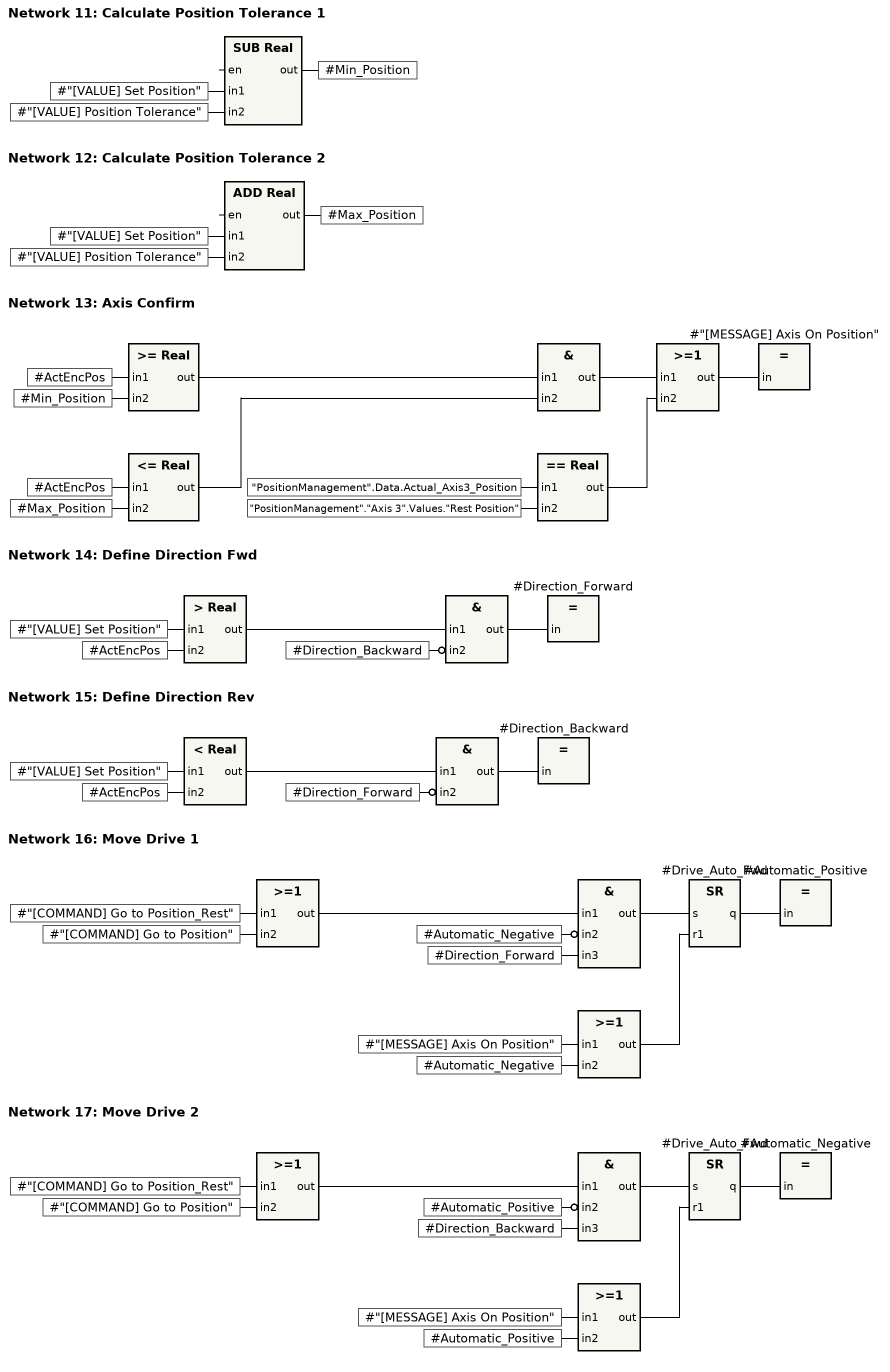
   #Min_Position := #"[VALUE] Set Position" - #"[VALUE] Position Tolerance";
END_REGION

REGION Network 12: Calculate Position Tolerance 2
   #Max_Position := #"[VALUE] Set Position" + #"[VALUE] Position Tolerance";
END_REGION

REGION Network 13: Axis Confirm
   #"[MESSAGE] Axis On Position" := ((#ActEncPos >= #Min_Position) AND (#ActEncPos <= #Max_Position)) OR ("PositionManagement".Data.Actual_Axis3_Position = "PositionManagement"."Axis 3".Values."Rest Position");
END_REGION

REGION Network 14: Define Direction Fwd
   #Direction_Forward := (#"[VALUE] Set Position" > #ActEncPos) AND NOT #Direction_Backward;
END_REGION

REGION Network 15: Define Direction Rev
   #Direction_Backward := (#"[VALUE] Set Position" < #ActEncPos) AND NOT #Direction_Forward;
END_REGION

REGION Network 16: Move Drive 1
   IF (#"[COMMAND] Go to Position_Rest" OR #"[COMMAND] Go to Position") AND NOT #Automatic_Negative AND #Direction_Forward THEN
       #Drive_Auto_Fwd := TRUE;   // SR flip-flop
   END_IF;
   IF #"[MESSAGE] Axis On Position" OR #Automatic_Negative THEN #Drive_Auto_Fwd := FALSE; END_IF;
   #Automatic_Positive := #Drive_Auto_Fwd;
END_REGION

REGION Network 17: Move Drive 2
   IF (#"[COMMAND] Go to Position_Rest" OR #"[COMMAND] Go to Position") AND NOT #Automatic_Positive AND #Direction_Backward THEN
       #Drive_Auto_Fwd := TRUE;   // SR flip-flop
   END_IF;
   IF #"[MESSAGE] Axis On Position" OR #Automatic_Positive THEN #Drive_Auto_Fwd := FALSE; END_IF;
   #Automatic_Negative := #Drive_Auto_Fwd;
END_REGION

REGION Network 18: Manual Displacement Positive
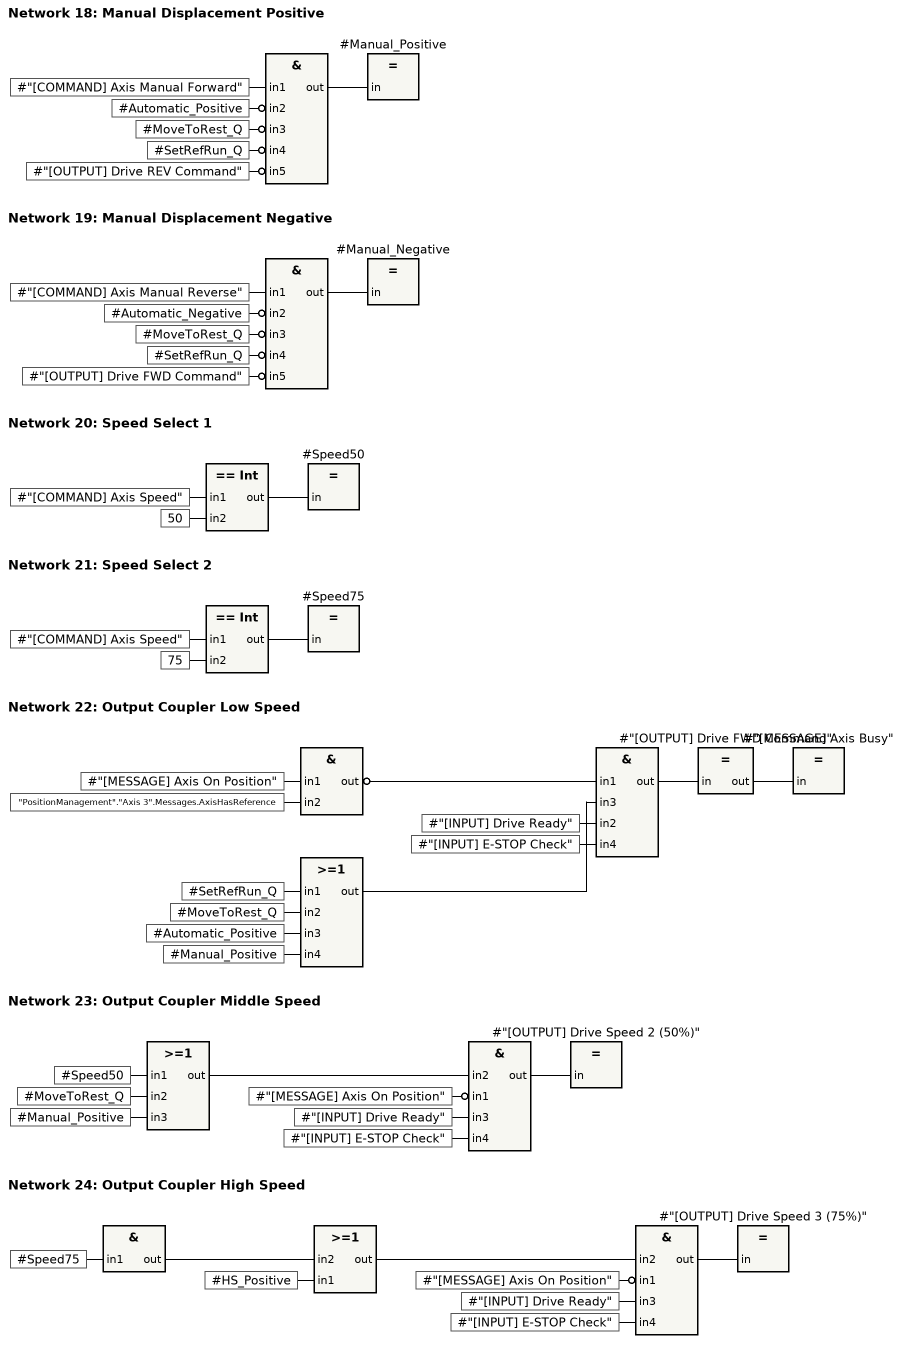
   #Manual_Positive := #"[COMMAND] Axis Manual Forward" AND NOT #Automatic_Positive AND NOT #MoveToRest_Q AND NOT #SetRefRun_Q AND NOT #"[OUTPUT] Drive REV Command";
END_REGION

REGION Network 19: Manual Displacement Negative
   #Manual_Negative := #"[COMMAND] Axis Manual Reverse" AND NOT #Automatic_Negative AND NOT #MoveToRest_Q AND NOT #SetRefRun_Q AND NOT #"[OUTPUT] Drive FWD Command";
END_REGION

REGION Network 20: Speed Select 1
   #Speed50 := #"[COMMAND] Axis Speed" = 50;
END_REGION

REGION Network 21: Speed Select 2
   #Speed75 := #"[COMMAND] Axis Speed" = 75;
END_REGION

REGION Network 22: Output Coupler Low Speed
   #_w1 := NOT (#"[MESSAGE] Axis On Position" AND "PositionManagement"."Axis 3".Messages.AxisHasReference) AND (#SetRefRun_Q OR #MoveToRest_Q OR #Automatic_Positive OR #Manual_Positive) AND #"[INPUT] Drive Ready" AND #"[INPUT] E-STOP Check";
   #"[OUTPUT] Drive FWD Command" := #_w1;
   #"[MESSAGE] Axis Busy" := #_w1;
END_REGION

REGION Network 23: Output Coupler Middle Speed
   #"[OUTPUT] Drive Speed 2 (50%)" := (#Speed50 OR #MoveToRest_Q OR #Manual_Positive) AND NOT #"[MESSAGE] Axis On Position" AND #"[INPUT] Drive Ready" AND #"[INPUT] E-STOP Check";
END_REGION

REGION Network 24: Output Coupler High Speed
   #"[OUTPUT] Drive Speed 3 (75%)" := (#Speed75 OR #HS_Positive) AND NOT #"[MESSAGE] Axis On Position" AND #"[INPUT] Drive Ready" AND #"[INPUT] E-STOP Check";
END_REGION

REGION Network 25: Output Coupler Reverse
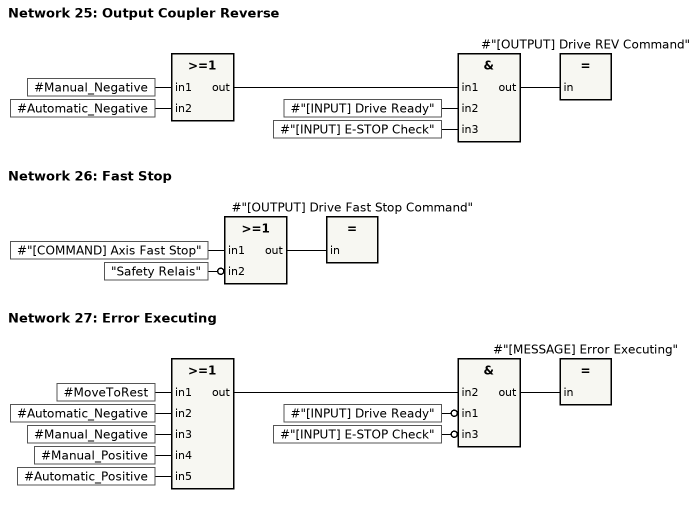
   #"[OUTPUT] Drive REV Command" := (#Manual_Negative OR #Automatic_Negative) AND #"[INPUT] Drive Ready" AND #"[INPUT] E-STOP Check";
END_REGION

REGION Network 26: Fast Stop
   #"[OUTPUT] Drive Fast Stop Command" := #"[COMMAND] Axis Fast Stop" OR NOT "Safety Relais";
END_REGION

REGION Network 27: Error Executing
   #"[MESSAGE] Error Executing" := (#MoveToRest OR #Automatic_Negative OR #Manual_Negative OR #Manual_Positive OR #Automatic_Positive) AND NOT #"[INPUT] Drive Ready" AND NOT #"[INPUT] E-STOP Check";
END_REGION
END_FUNCTION

(* ===== HMI "HMI_RT_2" =====
system functions are stored by id; their names below are inferred from use
connection "HMI_Connection_1": ETHERNET, SIMATIC S7 300/400 MPI

HMI tags "Default tag table"
   "Tag_ScreenNumber" : UInt, internal
   "Alle uitgangen(1)" : Bool = PLC "Alle uitgangen(1)" AT %I1.4, 1 s
   "Product op de band" : Bool = PLC "Sensor Op Band" AT %I0.6, 1 s
   "Product op de band(1)" : Bool = PLC "Sensor Op Band" AT %I0.6, 1 s
   "Trechter moet worden bijgevuld" : Bool = PLC "Sensor Trechter" AT %I0.5, 1 s
   "Voorverdeelwals staat in positie" : Bool = PLC "Sensor Wals (Option)" AT %I0.7, 1 s
   "Programma 1 draaid" : Bool = PLC "Programma 1" AT %I2.0, 1 s
   "Programma 2 draaid" : Bool = PLC "Programma 2" AT %I2.1, 1 s
   "Progrmma 3 draaid" : Bool = PLC "Programma 3" AT %I2.2, 1 s
   "Machine staat aan" : Bool = PLC "Start Machine" AT %I2.4, 1 s
   "Machine staat ui" : Bool = PLC "Stop Machine" AT %I2.5, 1 s
   "Noodstop machine" : Bool = PLC "ESB Pressend" AT %I1.1, 1 s
   "Startknop_Scherm" : Bool = PLC Startknop_Scherm AT %M15.0, 1 s
   "Stopknop_Scherm" : Bool = PLC Stopknop_Scherm AT %M15.1, 1 s
   "Systeem RUN" : Bool = PLC "Systeem RUN" AT %M0.0, 1 s
   "Reset Active" : Bool = PLC "Reset Active" AT %I1.2, 1 s
   "Drive 1 Ready" : Bool = PLC "Drive 1 Ready" AT %I0.0, 1 s
   "Drive 2 Ready" : Bool = PLC "Drive 2 Ready" AT %I0.1, 1 s
   "Drive 3 Ready" : Bool = PLC "Drive 3 Ready" AT %I0.2, 1 s
   "Drive 4 Ready" : Bool = PLC "Drive 4 Ready" AT %I0.3, 1 s
   "Drive 5 Ready" : Bool = PLC "Drive 5 Ready" AT %I0.4, 1 s
   "Drive 2 RUN FWD" : Bool = PLC "Drive 2 RUN FWD" AT %Q1.5, 1 s
   "Drive 1 RUN FWD" : Bool = PLC "Drive 1 RUN FWD" AT %Q1.0, 1 s
   "Drive 1 Speed 1" : Bool = PLC "Drive 1 Speed 1" AT %Q1.2, 1 s
   "Drive 1 Speed 2" : Bool = PLC "Drive 1 Speed 2" AT %Q1.3, 1 s
   "Drive 3 RUN FWD" : Bool = PLC "Drive 3 RUN FWD" AT %Q2.2, 1 s
   "Valve 1" : Bool = PLC "Valve 1" AT %Q4.6, 1 s
   "Drive 4 RUN FWD" : Bool = PLC "Drive 4 RUN FWD" AT %Q2.7, 1 s
   "StopAll" : Bool = PLC StopAll AT %M20.4, 1 s
   "Safety Relais" : Bool = PLC "Safety Relais" AT %Q0.0, 1 s
   "Drive_1_Manual" : Bool = PLC Drive_1_Manual AT %M50.1, 1 s
   "Stop_drive_1" : Bool = PLC Stop_drive_1 AT %M52.4, 1 s
   "Drive_2_Manual" : Bool = PLC Drive_2_Manual AT %M50.3, 1 s
   "Stop_drive_2" : Bool = PLC Stop_drive_2 AT %M52.5, 1 s
   "Drive_3_Manual" : Bool = PLC Drive_3_Manual AT %M50.5, 1 s
   "Stop_drive_3" : Bool = PLC Stop_drive_3 AT %M52.6, 1 s
   "Valve_1_Manual" : Bool = PLC Valve_1_Manual AT %M51.3, 1 s
   "Drive_4_Manual" : Bool = PLC Drive_4_Manual AT %M50.7, 1 s
   "Drive_5_Manual" : Bool = PLC Drive_5_Manual AT %M51.1, 1 s
   "Trechter_Bijvullen_Signaal" : Bool = PLC Trechter_Bijvullen_Signaal AT %M53.6, 1 s
   "RUN_Manual" : Bool = PLC RUN_Manual AT %M101.0, 1 s
   "Safety_Override" : Bool = PLC Safety_Override AT %M100.6, 1 s
   "Invert_Trechter_Sensor" : Bool = PLC Invert_Trechter_Sensor AT %M101.2, 1 s
   "Drive 1 REV]" : Bool = PLC "Drive 1 REV]" AT %Q1.1, 1 s
   "Drive 1 Rapid Stop" : Bool = PLC "Drive 1 Rapid Stop" AT %Q0.3, 1 s
   "Drive 2 Rapid Stop" : Bool = PLC "Drive 2 Rapid Stop" AT %Q0.4, 1 s
   "Drive 2 REV" : Bool = PLC "Drive 2 REV" AT %Q1.6, 1 s
   "Drive 3 Rapid Stop" : Bool = PLC "Drive 3 Rapid Stop" AT %Q0.5, 1 s
   "Drive 3 REV" : Bool = PLC "Drive 3 REV" AT %Q2.3, 1 s
   "Disable_Module" : Bool = PLC Disable_Module AT %M101.4, 1 s
   "PLCMemory_Safety_Delay" : Time = PLC PLCMemory.Safety_Delay AT %DB15.DBD8, 1 s
   "PLCMemory_Magazijn_Sensor_Delay" : Time = PLC PLCMemory.Offset_Timers.Magazijn_Sensor_Delay AT %DB15.DBD600, 1 s
   "PLCMemory_Homing_Sensor_Wals_Offset_Test" : Time = PLC PLCMemory.Homing_Sensor_Wals_Offset_Test AT %DB15.DBD0, 1 s
   "PLCMemory_Wals_Delay_Offset" : Time = PLC PLCMemory.Wals_Delay_Offset AT %DB15.DBD4, 1 s
   "PLCMemory_Aanvoer_Start_Offset" : Time = PLC PLCMemory.Offset_Timers.Aanvoer_Start_Offset AT %DB15.DBD596, 1 s
   "PLCMemory_Aanvoer_Stop_Offset" : Time = PLC PLCMemory.Offset_Timers.Aanvoer_Stop_Offset AT %DB15.DBD604, 1 s
   "PLCMemory_Trilgoten_Start_Offset" : Time = PLC PLCMemory.Offset_Timers.Trilgoten_Start_Offset AT %DB15.DBD588, 1 s
   "PLCMemory_Trilgoten_Stop_Offset" : Time = PLC PLCMemory.Offset_Timers.Trilgoten_Stop_Offset AT %DB15.DBD592, 1 s
   "Alarm_Axis_Not_Position" : Bool = PLC Alarm_Axis_Not_Position AT %M54.1, 1 s
   "PLCMemory_WalsCheck_Time" : Time = PLC PLCMemory.WalsCheck_Time AT %DB15.DBD12, 1 s
   "Alarm_Product_Not_Position" : Bool = PLC Alarm_Product_Not_Position AT %M54.2, 1 s
   "PLCMemory_ProductCheck_Time" : Time = PLC PLCMemory.ProductCheck_Time AT %DB15.DBD16, 1 s
   "LED Programma 1" : Bool = PLC "LED Programma 1" AT %Q4.1, 1 s
   "LED Programma 2" : Bool = PLC "LED Programma 2" AT %Q4.2, 1 s
   "LED Programma 3" : Bool = PLC "LED Programma 3" AT %Q4.3, 1 s
   "PLCMemory_ProductIntervalTime" : Time = PLC PLCMemory.ProductIntervalTime AT %DB15.DBD20, 1 s
   "PLCMemory_TD_Products_Counter" : Int = PLC PLCMemory.TD_Products_Counter AT %DB15.DBW32, 1 s
   "ResetTotalProducts" : Bool = PLC ResetTotalProducts AT %M102.7, 1 s
   "Door_Safety_Alarm" : Bool = PLC Door_Safety_Alarm AT %M54.3, 1 s
   "ESB_Safety_Alarm" : Bool = PLC ESB_Safety_Alarm AT %M54.4, 1 s
   "Valve_2_Manual" : Bool = PLC Valve_2_Manual AT %M51.5, 1 s
   "Valve 2" : Bool = PLC "Valve 2" AT %Q4.7, 1 s
   "Cilinder Trechterwissel in" : Bool = PLC "Spare(5)" AT %I3.0, 1 s
   "Cilinder Trechterwissel uit" : Bool = PLC "Spare(6)" AT %I3.1, 1 s
   "Valve 3" : Bool = PLC "Valve 3" AT %Q5.0, 1 s
   "Valve 4" : Bool = PLC "Valve 4" AT %Q5.1, 1 s
   "Valve 5" : Bool = PLC "Valve 5" AT %Q5.2, 1 s
   "Valve_3_Manual" : Bool = PLC Valve_3_Manual AT %M51.7, 1 s
   "Valve_4_Manual" : Bool = PLC Valve_4_Manual AT %M52.1, 1 s
   "Valve_5_Manual" : Bool = PLC Valve_5_Manual AT %M52.3, 1 s
   "Drive 5 REV" : Bool = PLC "Drive 5 REV" AT %Q3.5, 1 s
   "Drive 5 RUN FWD" : Bool = PLC "Drive 5 RUN FWD" AT %Q3.4, 1 s
   "Drive 5 Rapid Stop" : Bool = PLC "Drive 5 Rapid Stop" AT %Q0.7, 1 s
   "ESB Oke" : Bool = PLC "ESB Oke" AT %I1.0, 1 s
   "Door 1 NC contact" : Bool = PLC "Door 1 NC contact" AT %I1.5, 1 s
   "Door 2 NC contact" : Bool = PLC "Door 2 NC contact" AT %I1.7, 1 s
   "Sensor_op_band_memory" : Bool = PLC Sensor_op_band_memory AT %M15.3, 1 s
   "Drive_3_Auto" : Bool = PLC Drive_3_Auto AT %M50.4, 1 s
   "WalsSensorMemory" : Bool = PLC WalsSensorMemory AT %M101.3, 1 s
   "Drive_2_Auto" : Bool = PLC Drive_2_Auto AT %M50.2, 1 s
   "Drive_1_Auto" : Bool = PLC Drive_1_Auto AT %M50.0, 1 s
   "Alarms_AlarmsWord" : Word = PLC Alarms.AlarmsWord AT %DB24.DBW2, 1 s
   "Clear_Error" : Int, internal
   "Alarms_AlarmStruct_Alarm_Drive1" : Bool = PLC Alarms.AlarmStruct.Alarm_Drive1 AT %DB24.DBX0.2, 1 s
   "Alarms_HMI_Alarm_Drive1" : Word = PLC Alarms.HMI_Alarm_Drive1 AT %DB24.DBW4, 1 s
   "Alarms_HMI_Alarm_Drive2" : Word = PLC Alarms.HMI_Alarm_Drive2 AT %DB24.DBW6, 1 s
   "Alarms_HMI_Alarm_Drive3" : Word = PLC Alarms.HMI_Alarm_Drive3 AT %DB24.DBW8, 1 s
   "Alarms_HMI_Alarm_Drive4" : Word = PLC Alarms.HMI_Alarm_Drive4 AT %DB24.DBW10, 1 s
   "Alarms_HMI_Alarm_Drive5" : Word = PLC Alarms.HMI_Alarm_Drive5 AT %DB24.DBW12, 1 s
   "Sleutelschakelaar_Ingang" : Bool = PLC "Noodsleutel(1)" AT %I1.3, 1 s
      on ChangeValue: function_a9b89908("PLCMemory_UsernameMemory", "PLCMemory_PasswordMemory")
   "PLCMemory_UsernameMemory" : String[254] = PLC PLCMemory.UsernameMemory AT %DB15.DBX34.0, 1 s
   "PLCMemory_PasswordMemory" : String[254] = PLC PLCMemory.PasswordMemory AT %DB15.DBX290.0, 1 s
   "Drive 4 REV" : Bool = PLC "Drive 4 REV" AT %Q3.0, 1 s
   "Drive 4 Rapid Stop" : Bool = PLC "Drive 4 Rapid Stop" AT %Q0.6, 1 s
   "PLCMemory_SpeedSettingsTakeover" : Bool = PLC PLCMemory.SpeedSettingsTakeover AT %DB15.DBX546.0, 1 s
   "PLCMemory_SpeedSettingBand" : Bool = PLC PLCMemory.SpeedSettingBand AT %DB15.DBX546.2, 1 s
   "PLCMemory_TimingSettingOvername" : Bool = PLC PLCMemory.TimingSettingOvername AT %DB15.DBX546.3, 1 s
   "PLCMemory_SpeedSettingOvername" : Bool = PLC PLCMemory.SpeedSettingOvername AT %DB15.DBX546.1, 1 s
   "PLCMemory_Overname_Start_Offset" : Time = PLC PLCMemory.Offset_Timers.Overname_Start_Offset AT %DB15.DBD608, 1 s
   "PLCMemory_Overname_Stop_Offset" : Time = PLC PLCMemory.Offset_Timers.Overname_Stop_Offset AT %DB15.DBD612, 1 s
   "PLCMemory_EncoderPosition" : Real = PLC PLCMemory.EncoderPosition AT %DB15.DBD548, 1 s
   "PLCMemory_StepSize" : Real = PLC PLCMemory.StepSize AT %DB15.DBD552, 1 s
   "PLCMemory_Desired_Encoder_Position" : Real = PLC PLCMemory.Desired_Encoder_Position AT %DB15.DBD556, 1 s
   "HMI_Des_Pos_Axis3" : Bool = PLC HMI_Des_Pos_Axis3 AT %M54.5, 1 s
   "PLCMemory_Encoder PulsOffset" : Time = PLC PLCMemory."Encoder PulsOffset" AT %DB15.DBD564, 1 s
   "PLCMemory_Tolerance" : Real = PLC PLCMemory.Tolerance AT %DB15.DBD560, 1 s
   "PLCMemory_Axis3_Ref_Pos" : Real = PLC PLCMemory.Axis3_Ref_Pos AT %DB15.DBD568, 1 s
   "Cleaning_Active" : Bool = PLC Cleaning_Active AT %M182.0, 1 s
   "Cleaning" : Bool = PLC Cleaning AT %I2.3, 1 s
   "Cleaning_Confirmed" : Bool = PLC Cleaning_Confirmed AT %M182.1, 1 s
   "Cleaning_Cancelled" : Bool = PLC Cleaning_Cancelled AT %M182.2, 1 s
   "Cleaning_Screen_Active" : Bool = PLC Cleaning_Screen_Active AT %M182.3, 1 s
   "Tag_19" : Bool = PLC Tag_19 AT %M160.0, 1 s
   "Safety_Doors" : Bool = PLC Safety_Doors AT %M112.2, 1 s
   "HMI_ManualControl" : Bool = PLC HMI_ManualControl AT %M182.5, 1 s
   "PositionManagement_Data_Actual_Axis1_Position" : Real = PLC PositionManagement.Data.Actual_Axis3_Position AT %DB51.DBD16, 100 ms
   "PositionManagement_Axis 3_Values_Set Position" : Real, internal
   "PositionManagement_Axis 3_Commands_Go To Position" : Bool = PLC PositionManagement."Axis 3".Commands."Go To Position" AT %DB51.DBX312.3, 1 s
   "PositionManagement_Axis 3_Values_Pulsfactor" : Real = PLC PositionManagement."Axis 3".Values.Pulsfactor AT %DB51.DBD306, 1 s
   "PositionManagement_Axis 3_Values_Position Offset" : Real = PLC PositionManagement."Axis 3".Values."Position Offset" AT %DB51.DBD302, 1 s
   "PositionManagement_Axis 3_Values_Reference Position" : Int = PLC PositionManagement."Axis 3".Values."Reference Position" AT %DB51.DBW280, 1 s
   "PositionManagement_Axis 3_Values_Rest Position" : Real = PLC PositionManagement."Axis 3".Values."Rest Position" AT %DB51.DBD286, 1 s
   "PositionManagement_Axis 3_Values_Axis Correction" : Real = PLC PositionManagement."Axis 3".Values."Axis Correction" AT %DB51.DBD298, 1 s
   "PositionManagement_Axis 3_Values_Axis_Speed" : Int = PLC PositionManagement."Axis 3".Values.Axis_Speed AT %DB51.DBW310, 1 s
   "Drive_3_Manual_Rev" : Bool = PLC Drive_3_Manual_Rev AT %M60.1, 1 s
   "Manual Jog Fwd" : Bool = PLC "Manual Jog Fwd" AT %M137.0, 1 s
   "Manual Jog Rev" : Bool = PLC "Manual Jog Rev" AT %M137.1, 1 s
   "Counter2_IW102" : Int = PLC Counter2_IW102 AT %IW102, 1 s
   "PositionManagement_Axis 3_Commands_Start Ref Run" : Bool = PLC PositionManagement."Axis 3".Commands."Start Ref Run" AT %DB51.DBX312.1, 1 s
   "PLCMemory_Disable_Modules_Disable_Aandruk1" : Bool = PLC PLCMemory.Disable_Modules.Disable_Aandruk1 AT %DB15.DBX586.3, 1 s
   "PLCMemory_Disable_Modules_Disable_Aandruk2" : Bool = PLC PLCMemory.Disable_Modules.Disable_Aandruk2 AT %DB15.DBX586.4, 1 s
   "PLCMemory_Disable_Modules_Disable_Aandruk3" : Bool = PLC PLCMemory.Disable_Modules.Disable_Aandruk3 AT %DB15.DBX586.5, 1 s
   "PLCMemory_Disable_Modules_Disable_Blaaspuls" : Bool = PLC PLCMemory.Disable_Modules.Disable_Blaaspuls AT %DB15.DBX586.6, 1 s
   "PLCMemory_Disable_Modules_Disable_Afsluiter" : Bool = PLC PLCMemory.Disable_Modules.Disable_Afsluiter AT %DB15.DBX587.0, 1 s
   "PLCMemory_Offset_Timers_BlowOff_CycleTime" : Time = PLC PLCMemory.Offset_Timers.BlowOff_CycleTime AT %DB15.DBD624, 1 s
   "PLCMemory_Offset_Timers_Blow_Off_PulseTime" : Time = PLC PLCMemory.Offset_Timers.Blow_Off_PulseTime AT %DB15.DBD628, 1 s
   "PLCMemory_Disable_Modules_Disable_Retourband" : Bool = PLC PLCMemory.Disable_Modules.Disable_Retourband AT %DB15.DBX586.7, 1 s
   "PLCMemory_ProductBuffer_ProductsCount" : Int = PLC PLCMemory.ProductBuffer.ProductsCount AT %DB15.DBW636, 1 s
   "PLCMemory_ProductBufferBehindWals_Product_Count" : Int = PLC PLCMemory.ProductBufferBehindWals.Product_Count AT %DB15.DBW646, 1 s
   "PLCMemory_ProductBuffer_MoveTrigger" : Bool = PLC PLCMemory.ProductBuffer.MoveTrigger AT %DB15.DBX638.0, 1 s
   "Drive_4_Auto" : Bool = PLC Drive_4_Auto AT %M50.6, 1 s
   "ProductBuffer_V2_DB_SensorInput" : Bool = PLC ProductBuffer_V2_DB.SensorInput AT %DB66.DBX0.0, 1 s
   "PLCMemory_ProductBuffer_InsertIndex" : Int = PLC PLCMemory.ProductBuffer.InsertIndex AT %DB15.DBW640, 1 s
   "PLCMemory_SystemTime" : Time = PLC PLCMemory.SystemTime AT %DB15.DBD582, 1 s
   "PLCMemory" : Bool, internal
   "ProductBuffer_V2_DB_TriggerMovement" : Bool = PLC ProductBuffer_V2_DB.TriggerMovement AT %DB66.DBX12.0, 1 s
   "ProductBuffer_V2_DB_TriggerFeedback" : Bool = PLC ProductBuffer_V2_DB.TriggerFeedback AT %DB66.DBX10.0, 1 s
   "ProductBuffer_V2_DB_StartTimes__0" : Time = PLC ProductBuffer_V2_DB.StartTimes._0 AT %DB66.DBD34, 1 s
   "ProductBuffer_V2_DB_StartTimes__1" : Time = PLC ProductBuffer_V2_DB.StartTimes._1 AT %DB66.DBD38, 1 s
   "ProductBuffer_V2_DB_StartTimes__2" : Time = PLC ProductBuffer_V2_DB.StartTimes._2 AT %DB66.DBD42, 1 s
   "ProductBuffer_V2_DB_StartTimes__3" : Time = PLC ProductBuffer_V2_DB.StartTimes._3 AT %DB66.DBD46, 1 s
   "ProductBuffer_V2_DB_StartTimes__4" : Time = PLC ProductBuffer_V2_DB.StartTimes._4 AT %DB66.DBD50, 1 s
   "ProductBuffer_V2_DB_StartTimes__5" : Time = PLC ProductBuffer_V2_DB.StartTimes._5 AT %DB66.DBD54, 1 s
   "ProductBuffer_V2_DB_StartTimes__6" : Time = PLC ProductBuffer_V2_DB.StartTimes._6 AT %DB66.DBD58, 1 s
   "ProductBuffer_V2_DB_StartTimes__7" : Time = PLC ProductBuffer_V2_DB.StartTimes._7 AT %DB66.DBD62, 1 s
   "ProductBuffer_V2_DB_StartTimes__8" : Time = PLC ProductBuffer_V2_DB.StartTimes._8 AT %DB66.DBD66, 1 s
   "ProductBuffer_V2_DB_StartTimes__9" : Time = PLC ProductBuffer_V2_DB.StartTimes._9 AT %DB66.DBD70, 1 s
   "ProductBuffer_V2_DB_Actives__0" : Bool = PLC ProductBuffer_V2_DB.Actives._0 AT %DB66.DBX74.0, 1 s
   "ProductBuffer_V2_DB_Actives__1" : Bool = PLC ProductBuffer_V2_DB.Actives._1 AT %DB66.DBX74.1, 1 s
   "ProductBuffer_V2_DB_Actives__3" : Bool = PLC ProductBuffer_V2_DB.Actives._3 AT %DB66.DBX74.3, 1 s
   "ProductBuffer_V2_DB_Actives__2" : Bool = PLC ProductBuffer_V2_DB.Actives._2 AT %DB66.DBX74.2, 1 s
   "ProductBuffer_V2_DB_Actives__4" : Bool = PLC ProductBuffer_V2_DB.Actives._4 AT %DB66.DBX74.4, 1 s
   "ProductBuffer_V2_DB_Actives__5" : Bool = PLC ProductBuffer_V2_DB.Actives._5 AT %DB66.DBX74.5, 1 s
   "ProductBuffer_V2_DB_Actives__6" : Bool = PLC ProductBuffer_V2_DB.Actives._6 AT %DB66.DBX74.6, 1 s
   "ProductBuffer_V2_DB_Actives__7" : Bool = PLC ProductBuffer_V2_DB.Actives._7 AT %DB66.DBX74.7, 1 s
   "ProductBuffer_V2_DB_Actives__8" : Bool = PLC ProductBuffer_V2_DB.Actives._8 AT %DB66.DBX75.0, 1 s
   "ProductBuffer_V2_DB_Actives__9" : Bool = PLC ProductBuffer_V2_DB.Actives._9 AT %DB66.DBX75.1, 1 s
   "ProductBuffer_V2_DB_Elapsed" : DInt = PLC ProductBuffer_V2_DB.Elapsed AT %DB66.DBD80, 100 ms
   "ProductBuffer_V2_DB_PrevSensor" : Bool = PLC ProductBuffer_V2_DB.PrevSensor AT %DB66.DBX76.0, 1 s
   "ProductBuffer_V2_DB_MovementActive" : Bool = PLC ProductBuffer_V2_DB.MovementActive AT %DB66.DBX76.1, 1 s
   "PLCMemory_ProductBuffer_DelayTime" : Time = PLC PLCMemory.ProductBuffer.DelayTime AT %DB15.DBD632, 1 s
   "PositionManagement_Demo_Pos_Desired_Pos" : Real = PLC PositionManagement.Demo_Pos.Desired_Pos AT %DB51.DBD1342, 1 s
   "PositionManagement_Demo_Pos_Start" : Bool = PLC PositionManagement.Demo_Pos.Start AT %DB51.DBX1346.0, 1 s
   "PositionManagement_Axis_1_Values_Reference Position" : Int = PLC PositionManagement.Axis_1.Values."Reference Position" AT %DB51.DBW1614, 1 s
   "EncoderBand_RawCounter" : Int = PLC EncoderBand_RawCounter AT %IW112, 1 s
   "EncoderBand_Alive" : Int = PLC EncoderBand_Alive AT %IW110, 1 s
   "PositionManagement_Axis_1_Values_Axis Correction" : Real = PLC PositionManagement.Axis_1.Values."Axis Correction" AT %DB51.DBD1632, 1 s
   "Zpuls_Encoder_Band" : Bool = PLC Zpuls_Encoder_Band AT %I110.3, 1 s
   "PositionManagement_Data_Actual_Axis1_Position(1)" : Real = PLC PositionManagement.Data.Actual_Axis1_Position AT %DB51.DBD20, 1 s

HMI tags "Tag table_1"
   "ProductNoPosition_Alarm" : Bool = PLC Alarm_Product_Not_Position AT %M54.2, 1 s
   "AlarmsWord" : Word = PLC Alarms.AlarmsWord AT %DB24.DBW2, 1 s
   "Show_Expl" : Bool, internal

discrete alarms
   1: 'Let op! Producten komen niet op positie!', class Errors, trigger "Alarms_AlarmsWord" bit 0
   2: 'Let op! Wals komt niet op positie!', class Errors, trigger "Alarms_AlarmsWord" bit 1
   3: 'Drive 1 krijgt geen voedingsspanning of gaat niet aan.', class Errors, trigger "Alarms_HMI_Alarm_Drive1" bit 0
   4: 'Drive 2 krijgt geen voedingsspanning of gaat niet aan.', class Errors, trigger "Alarms_HMI_Alarm_Drive2" bit 0
   5: 'Drive 3 krijgt geen voedingsspanning of gaat niet aan.', class Errors, trigger "Alarms_HMI_Alarm_Drive3" bit 0
   6: 'Drive 4 krijgt geen voedingsspanning of gaat niet aan.', class Errors, trigger "Alarms_HMI_Alarm_Drive4" bit 0
   7: 'Drive 5 krijgt geen voedingsspanning of gaat niet aan.', class Errors, trigger "Alarms_HMI_Alarm_Drive5" bit 0

text list "List_Deactivate_Module": 0 'False'; 0 'False'; 1 'True'

text list "SpeedSettingOvername": 0..1 'Linked to Drive 1'; 0 'Speed 1'; 1 'Speed 2'

text list "SpeedSettings": 0 'No'; 1 'Yes'; 2 'Yes'

text list "SpeedSettingBand": 0..1 'Speed 1'; 0 'Speed 1'; 1 'Speed 2'

text list "Enable / Disable List": 0 '√'; 0 '√'; 1 'x'

graphic list "Enable_Graphic": 0 'vink groen'; 1 'cross red'; 0 'vink groen'

Template "Template_1" 800x480
   SymbolicIOField "Symbolic_IO_Field_Screen" at 93,9 size 600x33; TextOff '0'; TextOn '1'; TextList "TextList_ScreenNames"
      ProcessValue <- "Tag_ScreenNumber"
      on Change: ActivateScreenByNumber("Tag_ScreenNumber", 0)
   DateTimeField "HmiScreenItemData" at 695,25 size 105x25
   DateTimeField "HmiScreenItemData_1" at 695,0 size 105x25
   GraphicView "Logo" at 0,0 size 91x51; Picture "Logo of HMI_1"

screen "Screen_Handbediening" 800x480, template "Popup_Parameters"
   on GenerateScreen: SetBit("HMI_ManualControl")
   on ClearScreen: ResetBit("HMI_ManualControl")
   Softkey "Softkey_F8" at 0,0 size 0x0
      on KeyDown: function_ee5b8808("Button_3")
      on KeyUp: function_f101fd67("Button_3")
   GraphicView "Graphic view_2" at 0,80 size 799x399; Picture "SketchupModel_EklundNotenmachine_WithSafety achtergrond HMI"
   Circle "Circle_1" at 263,287 size 18x18
      Appearance <- "Product op de band"
   Circle "Circle_2" at 319,130 size 18x18
      Appearance <- "Trechter moet worden bijgevuld"
   Circle "Circle_3" at 325,228 size 18x18
      Appearance <- "Voorverdeelwals staat in positie"
   Rectangle "Rectangle_2" at 671,126 size 74x19
      Appearance <- "Safety Relais"
   DateTimeField "Date/time field_1" at 6,447 size 313x31
   GraphicView "Graphic view_1" at 2,80 size 141x101; Picture "logoeklund"
   Button "Button_2" at 595,93 size 200x55; TextOff 'Invoer'
      on Click: ActivateScreen("Screen_Band", 0)
   Button "Button_4" at 595,158 size 200x55; TextOff 'Trilgoten'
      on Click: ActivateScreen("Screen_Trilgoten", 0)
   Button "Button_5" at 595,222 size 200x55; TextOff 'Doseerwals'
      on Click: ActivateScreen("Screen_Doseerwals", 0)
   Button "Button_7" at 595,349 size 200x55; TextOff 'Afdichtingssysteem'
      on Click: ActivateScreen("Screen_Afdichting", 0)
   Button "Button_9" at 595,285 size 200x55; TextOff 'Aanvoerwals'
      on Click: ActivateScreen("Screen_AanvoerWals", 0)
   Button "Button_10" at 595,414 size 200x55; TextOff 'Aandruksysteem'
      on Click: ActivateScreen("Screen_Aandrukken", 0)
   Button "Button_3" at 6,174 size 130x60; TextOff 'Startscherm'; TextOn 'Onderweg na vorig scherm'
      on Click: ActivateScreen("Start_Screen", 0); ResetBit("HMI_ManualControl")
   Button "Button_1" at 6,247 size 130x55; TextOff 'Safety I/O'
      on Click: ActivateScreen("Screen_Safety_I/O", 0)
   Button "Button_8" at 7,315 size 130x55; TextOff 'Settings'; Authorization "TD ELKUND"
      on Click: ActivateScreen("Screen_Settings", 0)
   Button "Button_6" at 7,382 size 130x55; TextOff 'Retoursysteem'
      on Click: ActivateScreen("Screen_RetourBand", 0)

screen "Start_Screen" 800x480, template "Popup_Parameters"
   GraphicView "Graphic view_1" at 0,89 size 799x390; Picture "SketchupModel_EklundNotenmachine_WithSafety achtergrond HMI"
   Button "Button_1" at 4,230 size 165x70; TextOff 'Handbediening'
      on Click: ActivateScreen("Screen_Handbediening", 0); SetBit("HMI_ManualControl")
   Circle "Circle_1" at 260,291 size 18x18
      Appearance <- "Product op de band"
   Circle "Circle_2" at 321,139 size 18x18
      Appearance <- "Trechter moet worden bijgevuld"
   Circle "Circle_3" at 323,230 size 18x18
      Appearance <- "Voorverdeelwals staat in positie"
   DateTimeField "Date/time field_1" at 4,193 size 179x31
   GraphicView "Graphic view_2" at 5,91 size 155x101; Picture "logoeklund"
   Button "Button_2" at 630,310 size 165x70; TextOff 'Touchscreen cal.'
      on Click: function_bc3e350c()
   Button "Button_3" at 630,390 size 165x70; TextOff 'Logs'
      on Click: ActivateScreen("AlarmWindow", 0)
   Button "Button_4" at 4,310 size 165x70; TextOff 'Automatiek'
      on Click: ActivateScreen("Screen_Automatiek", 0)
   Button "Button_5" at 630,230 size 165x70; TextOff 'Producten'
   Circle "Circle_4" at 667,146 size 18x18
      Appearance <- "Safety_Doors"
   Circle "Circle_5" at 667,128 size 18x18
      Appearance <- "Safety Relais"
   Rectangle "Rectangle_1" at 242,203 size 417x173
      Visibility <- "Cleaning_Screen_Active"
   TextField "Text field_1" at 331,214 size 241x23; Text 'Cleaning Stand Geactiveerd!'
      Visibility <- "Cleaning_Screen_Active"
   TextField "Text field_2" at 259,252 size 378x61; Text 'Let op! Maak trechter eerst zo leeg mogelijk, en klik dan pas op ja! Bij op JA klikken gaan alle assen bewegen.'
      Visibility <- "Cleaning_Screen_Active"
   Button "Clean_NoButton" at 475,327 size 78x41; TextOff 'Nee'
      on Click: SetBit("Cleaning_Cancelled")
      Visibility <- "Cleaning_Screen_Active"
   Button "Clean_YesButton" at 568,327 size 78x41; TextOff 'Ja'
      on Click: SetBit("Cleaning_Confirmed")
      Visibility <- "Cleaning_Screen_Active"
   GraphicView "Graphic view_3" at 618,206 size 37x37; Picture "Graphic_31"
      Visibility <- "Cleaning_Screen_Active"
   GraphicView "Graphic view_4" at 246,206 size 37x37; Picture "Graphic_31"
      Visibility <- "Cleaning_Screen_Active"

screen "IOScreen" 800x480
   TextField "Text field_1" at 30,20 size 37x23; Text 'I0.0'
      Appearance <- "Drive 1 Ready"
   TextField "Text field_2" at 30,40 size 37x23; Text 'I0.1'
      Appearance <- "Drive 2 Ready"
   TextField "Text field_3" at 30,60 size 37x23; Text 'I0.2'
      Appearance <- "Drive 3 Ready"
   TextField "Text field_4" at 30,80 size 37x23; Text 'I0.3'
      Appearance <- "Drive 4 Ready"
   TextField "Text field_5" at 30,100 size 37x23; Text 'I0.4'
      Appearance <- "Drive 5 Ready"
   TextField "Text field_6" at 30,120 size 37x23; Text 'I0.5'
      Appearance <- "Trechter moet worden bijgevuld"
   Button "Button_7" at 697,6 size 96x32; TextOff 'Home'
      on Click: ActivateScreen("Screen_Handbediening", 0)
   Softkey "Softkey_F1" at 0,0 size 0x0
      on KeyDown: function_ee5b8808("Button_7")
      on KeyUp: function_f101fd67("Button_7")

screen "Screen_Trilgoten" 800x480, template "Popup_Parameters_Manual"
   TextField "Text field_1" at 10,228 size 207x23; Text 'Handbediening Trilgoten'
   TextField "Text field_8" at 85,262 size 42x23; Text 'Rust'
      Visibility <- "Drive 2 RUN FWD"
   TextField "Text field_9" at 103,262 size 147x23; Text 'Trilgoten running'
      Visibility <- "Drive 2 RUN FWD"
   TextField "Text field_4" at 433,173 size 105x23; Text 'Drive Status'
   TextField "Text field_5" at 615,174 size 74x23; Text 'Not ready'
      Visibility <- "Drive 2 Ready"
   TextField "Text field_6" at 433,227 size 153x23; Text 'Start Timer motor'
   IOField "StartMotorTimer" at 614,223 size 96x32; FormatPattern 9999
      ProcessValue <- "PLCMemory_Trilgoten_Start_Offset"
   TextField "Text field_12" at 433,261 size 149x23; Text 'Stop Timer motor'
   IOField "I/O field_2" at 614,258 size 96x32; FormatPattern 9999
      ProcessValue <- "PLCMemory_Trilgoten_Stop_Offset"
   TextField "Template_Text field_1" at 433,140 size 197x23; Text 'Trilgoten - Parameters'
   Button "Button_5" at 25,306 size 135x70; TextOff 'Start FWD'
      on Click: SetBit("Drive_2_Manual")
      Appearance <- "Drive_2_Manual"
   Button "Button_6" at 205,306 size 135x70; TextOff 'Stop FWD'
      on Click: ResetBit("Drive_2_Manual")
   TextField "Text field_2" at 612,174 size 48x23; Text 'Ready'
      Visibility <- "Drive 2 Ready"
   Button "Button_1" at 25,390 size 135x70; TextOff 'Start Rev'
      on Click: SetBit("Drive 2 REV")
      Appearance <- "Drive 2 REV"
   Button "Button_2" at 205,390 size 135x70; TextOff 'Stop Rev'
      on Click: ResetBit("Drive 2 REV")
   GraphicView "Graphic view_1" at 252,136 size 133x112; Picture "MotoriconArrowLeftRight"
   Circle "Circle_1" at 255,180 size 20x20
      Appearance <- "Drive 2 REV"
   Circle "Circle_2" at 359,180 size 20x20
      Appearance <- "Drive 2 RUN FWD"
   Circle "Circle_3" at 616,197 size 20x20
      Appearance <- "Drive 2 Rapid Stop"
   TextField "Text field_3" at 433,198 size 101x23; Text 'Drive Brake'
   TextField "Text field_11" at 721,226 size 25x22; Text 'ms'
   TextField "Text field_7" at 720,262 size 25x22; Text 'ms'

screen "Screen_Band" 800x480, template "Popup_Parameters_Manual"
   on GenerateScreen: SetBit("HMI_ManualControl")
   on ClearScreen: ResetBit("HMI_ManualControl")
   TextField "Text field_5" at 581,180 size 48x23; Text 'Ready'
      Visibility <- "Drive 1 Ready"
   TextField "Text field_4" at 584,180 size 74x23; Text 'Not ready'
      Visibility <- "Drive 1 Ready"
   TextField "Template_Text field_1" at 423,141 size 230x23; Text 'Aanvoerband - Parameters'
   TextField "Text field_1" at 8,220 size 173x23; Text 'Handbediening Band'
   TextField "Text field_8" at 85,261 size 42x23; Text 'Rust'
      Visibility <- "Drive 1 Ready"
   TextField "Text field_9" at 103,261 size 113x23; Text 'Band running'
      Visibility <- "Drive 1 Ready"
   TextField "Text field_3" at 425,180 size 105x23; Text 'Drive Status'
   Button "Button_1" at 25,306 size 135x70; TextOff 'Start FWD'
      on Click: SetBit("Drive_1_Manual")
      Appearance <- "Drive_1_Manual"
   Button "Button_2" at 205,306 size 135x70; TextOff 'Stop FWD'
      on Click: ResetBit("Drive_1_Manual")
   Button "Button_5" at 25,390 size 135x70; TextOff 'Start Rev'
      on Click: SetBit("Drive 1 REV]")
      Appearance <- "Drive 1 REV]"
   Button "Button_6" at 205,390 size 135x70; TextOff 'Stop Rev'
      on Click: ResetBit("Drive 1 REV]")
   Group "Group" at 581,180 size 77x23
   GraphicView "Graphic view_1" at 202,133 size 179x113; Picture "MotoriconArrowLeftRight"
   Circle "Circle_1" at 218,176 size 20x20
      Appearance <- "Drive 1 REV]"
   Circle "Circle_2" at 344,176 size 20x20
      Appearance <- "Drive 1 RUN FWD"
   IOField "I/O field_1" at 623,227 size 96x32; FormatPattern 99999
      ProcessValue <- "PLCMemory_ProductIntervalTime"
   TextField "Text field_10" at 425,234 size 144x23; Text 'Product Interval:'
   TextField "Text field_11" at 727,231 size 25x22; Text 'ms'
   TextField "Text field_15" at 428,272 size 125x23; Text 'Speed settings'
   SymbolicIOField "Symbolic I/O field_2" at 624,267 size 117x32; TextOn '1'; TextOff '0'; TextList "SpeedSettingBand"; HelpText 'Choose the speedsettings for Drive 1. (Speed 1 default speed, Speed 2 is faster movement)'
      ProcessValue <- "PLCMemory_SpeedSettingBand"
      on Activate: InvertBit("Show_Expl")
      on Deactivate: InvertBit("Show_Expl")
      on Change: ResetBit("Show_Expl")
   TextField "Text field_6" at 429,354 size 165x23; Text 'Reference Position:'
   IOField "StartMotorTimer" at 625,350 size 96x32; FormatPattern 9999
      ProcessValue <- "PositionManagement_Axis_1_Values_Reference Position"
   TextField "Text field_12" at 430,395 size 116x23; Text 'Encoder Alive'
   IOField "I/O field_2" at 624,392 size 96x32; FormatPattern 99999
      ProcessValue <- "EncoderBand_Alive"
   Circle "Circle_3" at 588,204 size 20x20
      Appearance <- "Zpuls_Encoder_Band"
   TextField "Text field_2" at 425,204 size 148x23; Text 'Reference Sensor'
   TextField "Text field_17" at 429,313 size 167x23; Text 'Position Correction:'
   IOField "I/O field_6" at 625,308 size 96x32; FormatPattern 9.99
      ProcessValue <- "PositionManagement_Axis_1_Values_Axis Correction"
   TextField "Text field_18" at 725,354 size 31x22; Text 'mm'
   TextField "Text field_19" at 725,315 size 31x22; Text 'mm'
   TextField "Text field_22" at 727,396 size 45x22; Text 'Pulses'
   TextField "Text field_7" at 430,431 size 92x23; Text 'Raw Value'
   IOField "I/O field_7" at 624,428 size 96x32; FormatPattern 999999
      ProcessValue <- "EncoderBand_RawCounter"
   TextField "Text field_23" at 727,432 size 45x22; Text 'Pulses'
   IOField "I/O field_3" at 230,259 size 110x29; FormatPattern 9999.9999
      ProcessValue <- "PositionManagement_Data_Actual_Axis1_Position(1)"
   TextField "Text field_13" at 347,263 size 31x22; Text 'mm'